
           //Erase the remaining element
           #INO_tMergeBuffer.rgtMessages[#INO_tMergeBuffer.dNumOfMessage - 1].dCodeEvent := 0;
           #INO_tMergeBuffer.rgtMessages[#INO_tMergeBuffer.dNumOfMessage - 1].strIdent := '';
           #INO_tMergeBuffer.rgtMessages[#INO_tMergeBuffer.dNumOfMessage - 1].dEvent1 := 0;
           #INO_tMergeBuffer.rgtMessages[#INO_tMergeBuffer.dNumOfMessage - 1].dEvent2 := 0;
           #INO_tMergeBuffer.rgtMessages[#INO_tMergeBuffer.dNumOfMessage - 1].dEvent3 := 0;
           #INO_tMergeBuffer.rgtMessages[#INO_tMergeBuffer.dNumOfMessage - 1].dEvent4 := 0;
           #INO_tMergeBuffer.rgtMessages[#INO_tMergeBuffer.dNumOfMessage - 1].dEvent5 := 0;
           #INO_tMergeBuffer.rgtMessages[#INO_tMergeBuffer.dNumOfMessage - 1].dEvent6 := 0;
           #INO_tMergeBuffer.rgtMessages[#INO_tMergeBuffer.dNumOfMessage - 1].dEvent7 := 0;
           #INO_tMergeBuffer.rgtMessages[#INO_tMergeBuffer.dNumOfMessage - 1].dEvent8 := 0;
           #INO_tMergeBuffer.rgtMessages[#INO_tMergeBuffer.dNumOfMessage - 1].dEvent9 := 0;
           #INO_tMergeBuffer.rgtMessages[#INO_tMergeBuffer.dNumOfMessage - 1].dEvent10 := 0;

           //Decrement the counter
           //
           #INO_tMergeBuffer.dNumOfMessage := #INO_tMergeBuffer.dNumOfMessage - 1;

       END_IF;


       #OUT_xDataAvailable := true;


   END_IF;
END_FUNCTION

// folder: 06_Output

FUNCTION "OutputTaskSlow" : Void   // FC11, LAD
{ S7_Optimized_Access := 'TRUE' }
VERSION : 0.1
   VAR_TEMP
      TMP_xSpareOFF : Bool;
   END_VAR
BEGIN

REGION Network 1 (SCL)
   #TMP_xSpareOFF := FALSE;


   "o.R195AP1.R251KA1.EncoderCommutation" :="FB_DigitizerManager_V1_00_IDB".OUTPUTS.xSelectEncoder1;
   "o.R195AP1.R251KA2.Jog" := "FB_DigitizerManager_V1_00_IDB".OUTPUTS.xEnableJog;
   "o.R195AP1.R252HL1.SafetiesON" :="Z200".tOutputs.xSafetiesON;

   "o.R195AP1.R251KA3.CpuASerSel":="Z200".tOutputs.xPLC1On;
   "o.R195AP1.R251KA4.CpuBSerSel" := "Z200".tOutputs.xPLC2On;

   "o.R195AP1.R252HL2.EnableCPUA" :="Z200".tOutputs.xPLC1On;
   "o.R195AP1.R252HL2.EnableCPUB" :="Z200".tOutputs.xPLC2On;


   "o.MCC1256B1_IDevice" := "FB_YCuts1_V1_00_IDB".OUT_tIDeviceData;
   "o.MCC1256B2_IDevice" := "FB_YCuts2_V1_00_IDB".OUT_tIDeviceData;


   "o.MCC1204_IDeviceToMarkers" := "FB_Markers_V1.00_IDB".OUT_tIDeviceData;

   "o.R195AP1.M216YV1.DigitizerRise/descentEncoder1" := "FB_Digitizer_1_V1_00_IDB".OUTPUTS.xDescentEncoder;
   "o.R195AP1.M216YV2.DigitizeRise/descentEncoder2" := "FB_Digitizer_2_V1_00_IDB".OUTPUTS.xDescentEncoder;
   "o.R195AP1.R429YV1.StartFillingPumpCuttingTank" := "FB_Oil_V1_00_IDB".OUTPUT.xTankFillCut;
   "o.R195AP1.M221YV2.UpperHolderControl" := "FB_Snaproll_V1_00_IDB".tOutputs.xContrastActivation;
   "o.R195AP1.M221YV1.BreakoutBarControl" := "FB_Snaproll_V1_00_IDB".tOutputs.xRiseSnap;

   "o.R195AP1.M221HL1.CutTrasversalBridge1" := "FB_Snaproll_V1_00_IDB".tOutputs.rgxHLCutDoneXC[0];
   "o.R195AP1.M221HL2.CutTrasversalBridge2" := "FB_Snaproll_V1_00_IDB".tOutputs.rgxHLCutDoneXC[1];
   "o.R195AP1.M221HL3.CutTrasversalBridge3" := "FB_Snaproll_V1_00_IDB".tOutputs.rgxHLCutDoneXC[2];


   "o.R195AP1.M212SB3.M212SB6.GlassRequestQlt" := "FB_ManInsp_V1_00_IDB".OUTPUT.rgxQualityButtonsLamp[0];






   "o_HSCOutput_Count2".swGate := "FB_Digitizer_1_V1_00_IDB".OUTPUTS.xCounterSWGate;
   "o_HSCOutput_Count3".swGate := "FB_Digitizer_2_V1_00_IDB".OUTPUTS.xCounterSWGate;
END_REGION
END_FUNCTION

FUNCTION "OutputTaskFast" : Void   // FC12, LAD
{ S7_Optimized_Access := 'TRUE' }
VERSION : 0.1
BEGIN

REGION Network 1 (SCL)
   "o.R195AP1.R252KA1.SCANNER.RiseBreakingBar" := "FB_ISRASNAP_V1_00_IDB".tOutputs.xSnap;
   "o.R195AP1.R252KA2.SCANNER.GlassToSQC" := "FB_ISRASNAP_V1_00_IDB".tOutputs.xSnapQlt;
   "o.R195AP1.A252KA3.SCANNER.NoGlassBreak" := "FB_ISRA5D_IDB".OUT_xGlassBreak;

   "o_HSCOutput_Count1" := "FB_TrackEncoder_V1_00_IDB".OUT_tHSCCount;
END_REGION
END_FUNCTION

FUNCTION "OutputTaskMedium" : Void   // FC13, LAD
{ S7_Optimized_Access := 'TRUE' }
VERSION : 0.1
BEGIN
END_FUNCTION

FUNCTION "Output_Z201_Idevice" : Void   // FC31, LAD
{ S7_Optimized_Access := 'TRUE' }
VERSION : 0.1
   VAR_TEMP
      TMP_xSpareOFF : Bool;
   END_VAR
BEGIN

REGION Network 1 (SCL)
   #TMP_xSpareOFF := FALSE;



   "FB_CommunicationZ300_V1.00_DB".OUT.Z200.tOUT_Mcc1201."xA47.7" := "Z201".tOutputs.xSafetiesON;

   "FB_CommunicationZ300_V1.00_DB".OUT.Z200.tOUT_Mcc1301."xE.A126.0" := "Z201".tOutputs.xHLResetAnomaly;

   //"o.CS4202.E406AP1.E547SB3.StartCleaningZ301" := "Check";
   //"o.CS4202.E406AP1.E547SB2.ResetAnomalyZ301" := "Check";
   //"o.CS4202.E406AP1.E547SB2.ResetAnomalyZ302" := "Check";
   //"o.CS4202.E406AP1.E547SB4.StopCleaningZ301" := "Check";

   "FB_CommunicationZ300_V1.00_DB".OUT.Z200.tOUT_Mcc1301."xE.A126.6" := "FB_BD_BreakPH_V1_00_IDB".OUTPUT.xSirenBreakAlarm OR"FB_BD_DigitizerPH_V1_00_IDB".OUTPUT.xSirenBreakAlarm ;
   "FB_CommunicationZ300_V1.00_DB".OUT.Z200.tOUT_Mcc1201."xA46.0" :=  "FB_BD_BreakPH_V1_00_IDB".OUTPUT.xLampBreakAlarm OR  "FB_BD_DigitizerPH_V1_00_IDB".OUTPUT.xLampBreakAlarm;


   "FB_CommunicationZ300_V1.00_DB".OUT.Z200.tOUT_Mcc1201."xA87.2" := "FB_DropConveyor_IDB".OUTPUT.xDescentDrop;
   "FB_CommunicationZ300_V1.00_DB".OUT.Z200.tOUT_Mcc1201."xA87.1" := "FB_DropConveyor_IDB".OUTPUT.xRiseDrop;
   "FB_CommunicationZ300_V1.00_DB".OUT.Z200.tOUT_Mcc1201."xA44.4" := true;
   "FB_CommunicationZ300_V1.00_DB".OUT.Z200.tOUT_Mcc1201."xA46.3" := "FB_DropConveyor_IDB".OUTPUT.xHLDoorOpen;
   "FB_CommunicationZ300_V1.00_DB".OUT.Z200.tOUT_Mcc1201."xA46.2" := "FB_DropConveyor_IDB".OUTPUT.xHLUpDownPushbutton;
   "FB_CommunicationZ300_V1.00_DB".OUT.Z200.tOUT_Mcc1201."xA46.5":= "FB_DropConveyor_IDB".OUTPUT.xHLDoorOpen;
   "FB_CommunicationZ300_V1.00_DB".OUT.Z200.tOUT_Mcc1201."xA46.6" := "FB_DropConveyor_IDB".OUTPUT.xHLUpDownPushbutton;

   "FB_CommunicationZ300_V1.00_DB".OUT.Z200.tOUT_Mcc1201."xA87.4" := "FB_BreakerM206_V1_00_IDB".OUTPUT.xBreakerRun;
   "FB_CommunicationZ300_V1.00_DB".OUT.Z200.tOUT_Mcc1201."xA44.0" := "FB_BreakerM206_V1_00_IDB".OUTPUT.xToScrapingUnderZ200;

   "FB_CommunicationZ300_V1.00_DB".OUT.Z200.tOUT_Mcc1201."xA86.0":="Z201".tOutputs.xRunFanM216;
   "FB_CommunicationZ300_V1.00_DB".OUT.Z200.tOUT_Mcc1201."xA87.6" := "Z201".tOutputs.xRunFanM209;
   "FB_CommunicationZ300_V1.00_DB".OUT.Z200.tOUT_Mcc1201."xA47.0" := "Z201".tOutputs.xHLchipBlowerM209On;

   "FB_CommunicationZ300_V1.00_DB".OUT.Z200.tOUT_Mcc1201."xA47.2" := "FB_BreakerM206_V1_00_IDB".OUTPUT.xHlScrapinglineReady;
   "FB_CommunicationZ300_V1.00_DB".OUT.Z200.tOUT_Mcc1201."xA47.3" := "FB_BreakerM206_V1_00_IDB".OUTPUT.xHlScrapinglineNotReady;
   "FB_CommunicationZ300_V1.00_DB".OUT.Z200.tOUT_Mcc1201."xA44.3" := "Z201".tOutputs.xHAAlarm;

   "FB_CommunicationZ300_V1.00_DB".OUT.Z200.tOUT_Mcc1201."xA45.0" := "FB_IO_EmergencyCuttingBridge_DB".OUT_xSnap;
   "FB_CommunicationZ300_V1.00_DB".OUT.Z200.tOUT_Mcc1201."xA45.3" := "FB_IO_EmergencyCuttingBridge_DB".OUT_xStartCutCycle;
END_REGION
END_FUNCTION

// folder: 07_ArrayScada

FUNCTION "SCADA_Mapping" : Void   // FC26, SCL
{ S7_Optimized_Access := 'TRUE' }
VERSION : 0.1
   VAR_TEMP
      TMP_dIndex : DInt;
   END_VAR
BEGIN


       //Move M201 HMR
       "DB_Conveyor_M201_HMI".tHMR.xManualCommandEnabled := "FB_Z200Conveyor_M201_IDB".tHMR.xManualCommandEnabled;
       "DB_Conveyor_M201_HMI".tHMR.dState := "FB_Z200Conveyor_M201_IDB".tHMR.dState;
       "DB_Conveyor_M201_HMI".tHMR.dSpeedFeedback := "FB_Z200Conveyor_M201_IDB".tHMR.dSpeedFeedback;
       "DB_Conveyor_M201_HMI".tHMR.tManCmd.xFdbkRunFw := "FB_Z200Conveyor_M201_IDB".tHMR.tManCmd.xFdbkRunFw;

       //Move M201 HMW
       "FB_Z200Conveyor_M201_IDB".tHMW.xEnableManualCommand := "DB_Conveyor_M201_HMI".tHMW.xEnableManualCommand;
       "FB_Z200Conveyor_M201_IDB".tHMW.tManCmd.xRunFw := "DB_Conveyor_M201_HMI".tHMW.tManCmd.xRunFw;
       "FB_Z200Conveyor_M201_IDB".tHMW.dCurrentLimit := "DB_Conveyor_M201_HMI".tHMW.dCurrentLimit;
       "FB_Z200Conveyor_M201_IDB".tHMW.dSpeedCorrection := "DB_Conveyor_M201_HMI".tHMW.dSpeedCorrection;

       //Move M201 ALM
       "DB_Conveyor_M201_HMI".tALM.tF :="FB_Z200Conveyor_M201_IDB".tALM.tF;
       "DB_Conveyor_M201_HMI".tALM.tS := "FB_Z200Conveyor_M201_IDB".tALM.tS;
       "DB_Conveyor_M201_HMI".tALM.tW := "FB_Z200Conveyor_M201_IDB".tALM.tW;

       //Move M204 HMR
       "DB_Conveyor_M204_HMI".tHMR.xManualCommandEnabled := "FB_Z200Conveyor_M204_IDB".tHMR.xManualCommandEnabled;
       "DB_Conveyor_M204_HMI".tHMR.dState := "FB_Z200Conveyor_M204_IDB".tHMR.dState;
       "DB_Conveyor_M204_HMI".tHMR.dSpeedFeedback := "FB_Z200Conveyor_M204_IDB".tHMR.dSpeedFeedback;
       "DB_Conveyor_M204_HMI".tHMR.tManCmd.xFdbkRunFw := "FB_Z200Conveyor_M204_IDB".tHMR.tManCmd.xFdbkRunFw;

       //Move M204 HMW
       "FB_Z200Conveyor_M204_IDB".tHMW.xEnableManualCommand := "DB_Conveyor_M204_HMI".tHMW.xEnableManualCommand;
       "FB_Z200Conveyor_M204_IDB".tHMW.tManCmd.xRunFw := "DB_Conveyor_M204_HMI".tHMW.tManCmd.xRunFw;
       "FB_Z200Conveyor_M204_IDB".tHMW.dCurrentLimit := "DB_Conveyor_M204_HMI".tHMW.dCurrentLimit;
       "FB_Z200Conveyor_M204_IDB".tHMW.dSpeedCorrection := "DB_Conveyor_M204_HMI".tHMW.dSpeedCorrection;

       //Move M204 ALM
       "DB_Conveyor_M204_HMI".tALM.tF := "FB_Z200Conveyor_M204_IDB".tALM.tF;
       "DB_Conveyor_M204_HMI".tALM.tS := "FB_Z200Conveyor_M204_IDB".tALM.tS;
       "DB_Conveyor_M204_HMI".tALM.tW := "FB_Z200Conveyor_M204_IDB".tALM.tW;

       //Move M205 HMR
       "DB_Conveyor_M205_HMI".tHMR.xManualCommandEnabled := "FB_Z200Conveyor_M205_IDB".tHMR.xManualCommandEnabled;
       "DB_Conveyor_M205_HMI".tHMR.dState := "FB_Z200Conveyor_M205_IDB".tHMR.dState;
       "DB_Conveyor_M205_HMI".tHMR.dSpeedFeedback := "FB_Z200Conveyor_M205_IDB".tHMR.dSpeedFeedback;
       "DB_Conveyor_M205_HMI".tHMR.tManCmd.xFdbkRunFw := "FB_Z200Conveyor_M205_IDB".tHMR.tManCmd.xFdbkRunFw;

       //Move M205 HMW
       "FB_Z200Conveyor_M205_IDB".tHMW.xEnableManualCommand := "DB_Conveyor_M205_HMI".tHMW.xEnableManualCommand;
       "FB_Z200Conveyor_M205_IDB".tHMW.tManCmd.xRunFw := "DB_Conveyor_M205_HMI".tHMW.tManCmd.xRunFw;
       "FB_Z200Conveyor_M205_IDB".tHMW.dCurrentLimit := "DB_Conveyor_M205_HMI".tHMW.dCurrentLimit;
       "FB_Z200Conveyor_M205_IDB".tHMW.dSpeedCorrection := "DB_Conveyor_M205_HMI".tHMW.dSpeedCorrection;

       //Move M205 ALM
       "DB_Conveyor_M205_HMI".tALM.tF := "FB_Z200Conveyor_M205_IDB".tALM.tF;


       //Move M208 HMR
       "DB_Conveyor_M208_HMI".tHMR.xManualCommandEnabled := "FB_Z200Conveyor_M208_IDB".tHMR.xManualCommandEnabled;
       "DB_Conveyor_M208_HMI".tHMR.dState := "FB_Z200Conveyor_M208_IDB".tHMR.dState;
       "DB_Conveyor_M208_HMI".tHMR.dSpeedFeedback := "FB_Z200Conveyor_M208_IDB".tHMR.dSpeedFeedback;
       "DB_Conveyor_M208_HMI".tHMR.tManCmd.xFdbkRunFw := "FB_Z200Conveyor_M208_IDB".tHMR.tManCmd.xFdbkRunFw;

       //Move M208 HMW
       "FB_Z200Conveyor_M208_IDB".tHMW.xEnableManualCommand := "DB_Conveyor_M208_HMI".tHMW.xEnableManualCommand;
       "FB_Z200Conveyor_M208_IDB".tHMW.tManCmd.xRunFw := "DB_Conveyor_M208_HMI".tHMW.tManCmd.xRunFw;
       "FB_Z200Conveyor_M208_IDB".tHMW.dCurrentLimit := "DB_Conveyor_M208_HMI".tHMW.dCurrentLimit;
       "FB_Z200Conveyor_M208_IDB".tHMW.dSpeedCorrection := "DB_Conveyor_M208_HMI".tHMW.dSpeedCorrection;

       //Move M208 ALM
       "DB_Conveyor_M208_HMI".tALM.tF := "FB_Z200Conveyor_M208_IDB".tALM.tF;
       "DB_Conveyor_M208_HMI".tALM.tS:= "FB_Z200Conveyor_M208_IDB".tALM.tS;
       "DB_Conveyor_M208_HMI".tALM.tW := "FB_Z200Conveyor_M208_IDB".tALM.tW;

        //Move M211 HMR
       "DB_Conveyor_M211_HMI".tHMR.xManualCommandEnabled := "FB_Z200Conveyor_M211_iDB".tHMR.xManualCommandEnabled;
       "DB_Conveyor_M211_HMI".tHMR.dState := "FB_Z200Conveyor_M211_iDB".tHMR.dState;
       "DB_Conveyor_M211_HMI".tHMR.dSpeedFeedback := "FB_Z200Conveyor_M211_iDB".tHMR.dSpeedFeedback;
       "DB_Conveyor_M211_HMI".tHMR.tManCmd.xFdbkRunFw := "FB_Z200Conveyor_M211_iDB".tHMR.tManCmd.xFdbkRunFw;

       //Move M211 HMW
       "FB_Z200Conveyor_M211_iDB".tHMW.xEnableManualCommand := "DB_Conveyor_M211_HMI".tHMW.xEnableManualCommand;
       "FB_Z200Conveyor_M211_iDB".tHMW.tManCmd.xRunFw := "DB_Conveyor_M211_HMI".tHMW.tManCmd.xRunFw;
       "FB_Z200Conveyor_M211_iDB".tHMW.dCurrentLimit := "DB_Conveyor_M211_HMI".tHMW.dCurrentLimit;
       "FB_Z200Conveyor_M211_iDB".tHMW.dSpeedCorrection := "DB_Conveyor_M211_HMI".tHMW.dSpeedCorrection;

       //Move M211 ALM
       "DB_Conveyor_M211_HMI".tALM.tF := "FB_Z200Conveyor_M211_iDB".tALM.tF;
       "DB_Conveyor_M211_HMI".tALM.tS := "FB_Z200Conveyor_M211_iDB".tALM.tS;
       "DB_Conveyor_M211_HMI".tALM.tW := "FB_Z200Conveyor_M211_iDB".tALM.tW;



       //Move M214 HMR
       "DB_Conveyor_M214_HMI".tHMR.xManualCommandEnabled := "FB_Z200Conveyor_M214_iDB".tHMR.xManualCommandEnabled;
       "DB_Conveyor_M214_HMI".tHMR.dState := "FB_Z200Conveyor_M214_iDB".tHMR.dState;
       "DB_Conveyor_M214_HMI".tHMR.dSpeedFeedback := "FB_Z200Conveyor_M214_iDB".tHMR.dSpeedFeedback;
       "DB_Conveyor_M214_HMI".tHMR.tManCmd.xFdbkRunFw := "FB_Z200Conveyor_M214_iDB".tHMR.tManCmd.xFdbkRunFw;

       //Move M214 HMW
       "FB_Z200Conveyor_M214_iDB".tHMW.xEnableManualCommand := "DB_Conveyor_M214_HMI".tHMW.xEnableManualCommand;
       "FB_Z200Conveyor_M214_iDB".tHMW.tManCmd.xRunFw := "DB_Conveyor_M214_HMI".tHMW.tManCmd.xRunFw;
       "FB_Z200Conveyor_M214_iDB".tHMW.dCurrentLimit := "DB_Conveyor_M214_HMI".tHMW.dCurrentLimit;
       "FB_Z200Conveyor_M214_iDB".tHMW.dSpeedCorrection := "DB_Conveyor_M214_HMI".tHMW.dSpeedCorrection;

       //Move M214 ALM
       "DB_Conveyor_M214_HMI".tALM.tF := "FB_Z200Conveyor_M214_iDB".tALM.tF;
       "DB_Conveyor_M214_HMI".tALM.tS := "FB_Z200Conveyor_M214_iDB".tALM.tS;
       "DB_Conveyor_M214_HMI".tALM.tW := "FB_Z200Conveyor_M214_iDB".tALM.tW;

       //Move M218 HMR
       "DB_Conveyor_M218_HMI".tHMR.xManualCommandEnabled := "FB_Z200Conveyor_M218_IDB".tHMR.xManualCommandEnabled;
       "DB_Conveyor_M218_HMI".tHMR.dState := "FB_Z200Conveyor_M218_IDB".tHMR.dState;
       "DB_Conveyor_M218_HMI".tHMR.dSpeedFeedback := "FB_Z200Conveyor_M218_IDB".tHMR.dSpeedFeedback;
       "DB_Conveyor_M218_HMI".tHMR.tManCmd.xFdbkRunFw := "FB_Z200Conveyor_M218_IDB".tHMR.tManCmd.xFdbkRunFw;

       //Move M218 HMW
       "FB_Z200Conveyor_M218_IDB".tHMW.xEnableManualCommand := "DB_Conveyor_M218_HMI".tHMW.xEnableManualCommand;
       "FB_Z200Conveyor_M218_IDB".tHMW.tManCmd.xRunFw := "DB_Conveyor_M218_HMI".tHMW.tManCmd.xRunFw;
       "FB_Z200Conveyor_M218_IDB".tHMW.dCurrentLimit := "DB_Conveyor_M218_HMI".tHMW.dCurrentLimit;
       "FB_Z200Conveyor_M218_IDB".tHMW.dSpeedCorrection := "DB_Conveyor_M218_HMI".tHMW.dSpeedCorrection;

       //Move M218 ALM
       "DB_Conveyor_M218_HMI".tALM.tF := "FB_Z200Conveyor_M218_IDB".tALM.tF;
       "DB_Conveyor_M218_HMI".tALM.tS := "FB_Z200Conveyor_M218_IDB".tALM.tS;
       "DB_Conveyor_M218_HMI".tALM.tW := "FB_Z200Conveyor_M218_IDB".tALM.tW;

       //Move M206 HMR
       "DB_Breaker_M206_HMI".tHMR.xSpare1 :="FB_BreakerM206_V1_00_IDB".tHMR.xEnabledRunAlwaysModeBreaker;
       "DB_Breaker_M206_HMI".tHMR.xManualCommandEnabled := "FB_BreakerM206_V1_00_IDB".tHMR.xManualCommandEnabled;
       "DB_Breaker_M206_HMI".tHMR.tManCmd.xRunFdbk := "FB_BreakerM206_V1_00_IDB".tHMR.tManCmd.xRunFdbk;

       //Move M206 HMW
       "FB_BreakerM206_V1_00_IDB".tHMW.dBreakerRetainTime_s := "DB_Breaker_M206_HMI".tHMW.dBreakerRetainTime_s;
       "FB_BreakerM206_V1_00_IDB".tHMW.xEnableManualCommand := "DB_Breaker_M206_HMI".tHMW.xEnableManualCommand;
       "FB_BreakerM206_V1_00_IDB".tHMW.xEnableRunAlwaysModeBreaker := "DB_Breaker_M206_HMI".tHMW.xEnableRunAlwaysModeBreaker;
       "FB_BreakerM206_V1_00_IDB".tHMW.tManCmd.xRun := "DB_Breaker_M206_HMI".tHMW.tManCmd.xRun;

       //Move M206 ALM 
       "DB_Breaker_M206_HMI".tALM.tF :="FB_BreakerM206_V1_00_IDB".tALM.tF;
       "DB_Breaker_M206_HMI".tALM.tS :="FB_BreakerM206_V1_00_IDB".tALM.tS;
       "DB_Breaker_M206_HMI".tALM.tW :="FB_BreakerM206_V1_00_IDB".tALM.tW;

       //Move MAN INSP HMR
       //
       "DB_MAN_INSP_HMI".tHMR.xManualCommandEnabled := "FB_ManInsp_V1_00_IDB".tHMR.xManComEn;
       "DB_MAN_INSP_HMI".tHMR.dDistanceSnaproll_cmm := "FB_ManInsp_V1_00_IDB".tHMR.dDistanceSnaproll_cmm;
       "DB_MAN_INSP_HMI".tHMR.tManCmd.xSpare1 := "FB_ManInsp_V1_00_IDB".tHMR.tManFdbk.xFanCommand; 

       //Move MAN INSP   HMW
       "FB_ManInsp_V1_00_IDB".tHMW.xUpdateDistanceSnaproll := "DB_MAN_INSP_HMI".tHMW.xUpdateDistanceSnaproll;
       "FB_ManInsp_V1_00_IDB".tHMW.xEnDisManCom := "DB_MAN_INSP_HMI".tHMW.xEnableManualCommand;
       "FB_ManInsp_V1_00_IDB".tHMW.rgxEnabledContinuosDef[0] := "DB_MAN_INSP_HMI".tHMW."xEnabledContinuosDef[0]";
       "FB_ManInsp_V1_00_IDB".tHMW.rgxEnabledContinuosDef[1] := "DB_MAN_INSP_HMI".tHMW."xEnabledContinuosDef[1]";
       "FB_ManInsp_V1_00_IDB".tHMW.rgxEnabledContinuosDef[2] := "DB_MAN_INSP_HMI".tHMW."xEnabledContinuosDef[2]";
       "FB_ManInsp_V1_00_IDB".tHMW.rgxEnabledContinuosDef[3] := "DB_MAN_INSP_HMI".tHMW."xEnabledContinuosDef[3]";
       "FB_ManInsp_V1_00_IDB".tHMW.tMan.xFanCommand := "DB_MAN_INSP_HMI".tHMW.tManCmd.xSpare0;


       //Move MAN INSP  ALM  
       "DB_MAN_INSP_HMI".tALM.tF := "FB_ManInsp_V1_00_IDB".tALM.tF;
       "DB_MAN_INSP_HMI".tALM.tS := "FB_ManInsp_V1_00_IDB".tALM.tS;
       "DB_MAN_INSP_HMI".tALM.tW := "FB_ManInsp_V1_00_IDB".tALM.tW;

       //Move BREAK DETECTOR HMR

       "DB_Break_detector_M202_HMI".tHMR."xPhotoStatus[0]" := "FB_BD_BreakPH_V1_00_IDB".tHMR.rgxPhotoStatus[0];
       "DB_Break_detector_M202_HMI".tHMR."xPhotoStatus[1]" := "FB_BD_BreakPH_V1_00_IDB".tHMR.rgxPhotoStatus[1];
       "DB_Break_detector_M202_HMI".tHMR."xPhotoStatus[2]" := "FB_BD_BreakPH_V1_00_IDB".tHMR.rgxPhotoStatus[2];
       "DB_Break_detector_M202_HMI".tHMR."xPhotoStatus[3]" := "FB_BD_BreakPH_V1_00_IDB".tHMR.rgxPhotoStatus[3];
       "DB_Break_detector_M202_HMI".tHMR."xPhotoStatus[4]" := "FB_BD_BreakPH_V1_00_IDB".tHMR.rgxPhotoStatus[4];
       "DB_Break_detector_M202_HMI".tHMR."xPhotoStatus[5]" := "FB_BD_BreakPH_V1_00_IDB".tHMR.rgxPhotoStatus[5];
       "DB_Break_detector_M202_HMI".tHMR."xPhotoStatus[6]" := "FB_BD_BreakPH_V1_00_IDB".tHMR.rgxPhotoStatus[6];
       "DB_Break_detector_M202_HMI".tHMR."xPhotoStatus[7]" := "FB_BD_BreakPH_V1_00_IDB".tHMR.rgxPhotoStatus[7];
       "DB_Break_detector_M202_HMI".tHMR."xPhotoStatus[8]" := "FB_BD_BreakPH_V1_00_IDB".tHMR.rgxPhotoStatus[8];
       "DB_Break_detector_M202_HMI".tHMR."xPhotoStatus[9]" := "FB_BD_BreakPH_V1_00_IDB".tHMR.rgxPhotoStatus[9];

       "DB_Break_detector_M202_HMI".tHMR.dDistanceSnaproll_cmm := "FB_BD_BreakPH_V1_00_IDB".tHMR.dDistanceSnaproll_cmm;
       "DB_Break_detector_M202_HMI".tHMR.dStatus := "FB_BD_BreakPH_V1_00_IDB".tHMR.dStatus;
       "DB_Break_detector_M202_HMI".tHMR."dPhotoAbilitation[0]" := "FB_BD_BreakPH_V1_00_IDB".tHMR.rgdPhotoAbilitation[0];
       "DB_Break_detector_M202_HMI".tHMR."dPhotoAbilitation[1]" := "FB_BD_BreakPH_V1_00_IDB".tHMR.rgdPhotoAbilitation[1];
       "DB_Break_detector_M202_HMI".tHMR."dPhotoAbilitation[2]" := "FB_BD_BreakPH_V1_00_IDB".tHMR.rgdPhotoAbilitation[2];
       "DB_Break_detector_M202_HMI".tHMR."dPhotoAbilitation[3]" := "FB_BD_BreakPH_V1_00_IDB".tHMR.rgdPhotoAbilitation[3];
       "DB_Break_detector_M202_HMI".tHMR."dPhotoAbilitation[4]" := "FB_BD_BreakPH_V1_00_IDB".tHMR.rgdPhotoAbilitation[4];
       "DB_Break_detector_M202_HMI".tHMR."dPhotoAbilitation[5]" := "FB_BD_BreakPH_V1_00_IDB".tHMR.rgdPhotoAbilitation[5];
       "DB_Break_detector_M202_HMI".tHMR."dPhotoAbilitation[6]" := "FB_BD_BreakPH_V1_00_IDB".tHMR.rgdPhotoAbilitation[6];
       "DB_Break_detector_M202_HMI".tHMR."dPhotoAbilitation[7]" := "FB_BD_BreakPH_V1_00_IDB".tHMR.rgdPhotoAbilitation[7];
       "DB_Break_detector_M202_HMI".tHMR."dPhotoAbilitation[8]" := "FB_BD_BreakPH_V1_00_IDB".tHMR.rgdPhotoAbilitation[8];
       "DB_Break_detector_M202_HMI".tHMR."dPhotoAbilitation[9]" := "FB_BD_BreakPH_V1_00_IDB".tHMR.rgdPhotoAbilitation[9];

       //Move BREAK DETECTOR HMW
       "FB_BD_BreakPH_V1_00_IDB".tHMW.xUpdateDistanceSnap := "DB_Break_detector_M202_HMI".tHMW.xUpdateDistanceSnaproll;

       "FB_BD_BreakPH_V1_00_IDB".tHMW.rgxEnabledPhotocell[0] := "DB_Break_detector_M202_HMI".tHMW."xPhotoEnabled[0]";
       "FB_BD_BreakPH_V1_00_IDB".tHMW.rgxEnabledPhotocell[1] := "DB_Break_detector_M202_HMI".tHMW."xPhotoEnabled[1]";
       "FB_BD_BreakPH_V1_00_IDB".tHMW.rgxEnabledPhotocell[2] := "DB_Break_detector_M202_HMI".tHMW."xPhotoEnabled[2]";
       "FB_BD_BreakPH_V1_00_IDB".tHMW.rgxEnabledPhotocell[3] := "DB_Break_detector_M202_HMI".tHMW."xPhotoEnabled[3]";
       "FB_BD_BreakPH_V1_00_IDB".tHMW.rgxEnabledPhotocell[4] := "DB_Break_detector_M202_HMI".tHMW."xPhotoEnabled[4]";
       "FB_BD_BreakPH_V1_00_IDB".tHMW.rgxEnabledPhotocell[5] := "DB_Break_detector_M202_HMI".tHMW."xPhotoEnabled[5]";
       "FB_BD_BreakPH_V1_00_IDB".tHMW.rgxEnabledPhotocell[6] := "DB_Break_detector_M202_HMI".tHMW."xPhotoEnabled[6]";
       "FB_BD_BreakPH_V1_00_IDB".tHMW.rgxEnabledPhotocell[7] := "DB_Break_detector_M202_HMI".tHMW."xPhotoEnabled[7]";
       "FB_BD_BreakPH_V1_00_IDB".tHMW.rgxEnabledPhotocell[8] := "DB_Break_detector_M202_HMI".tHMW."xPhotoEnabled[8]";
       "FB_BD_BreakPH_V1_00_IDB".tHMW.rgxEnabledPhotocell[9] := "DB_Break_detector_M202_HMI".tHMW."xPhotoEnabled[9]";

       "FB_BD_BreakPH_V1_00_IDB".tHMW.dDistanceSnaproll_cmm := "DB_Break_detector_M202_HMI".tHMW.dDistanceSnaproll_cmm;
       "FB_BD_BreakPH_V1_00_IDB".tHMW.dMinBreakSize_cmm :="DB_Break_detector_M202_HMI".tHMW.dMinBreakSize_cmm;

       //Move BREAK DETECTOR ALM
       "DB_Break_detector_M202_HMI".tALM.tF := "FB_BD_BreakPH_V1_00_IDB".tALM.tF;
       "DB_Break_detector_M202_HMI".tALM.tS := "FB_BD_BreakPH_V1_00_IDB".tALM.tS;
       "DB_Break_detector_M202_HMI".tALM.tW := "FB_BD_BreakPH_V1_00_IDB".tALM.tW;

       //Move ISRA HMR
       "DB_ISRA_HMI".tHMR.xScannerON := "FB_ISRA5D_IDB".tHMR.xScannerON;

       "DB_ISRA_HMI".tHMR.dCurrentGrossWander_cmm := "FB_ISRA5D_IDB".tHMR.dCurrentGrossWander_cmm;
       "DB_ISRA_HMI".tHMR.dCurrentGrossWidth_cmm := "FB_ISRA5D_IDB".tHMR.dCurrentGrossWidth_cmm;
       "DB_ISRA_HMI".tHMR.dCurrentNetWander_cmm := "FB_ISRA5D_IDB".tHMR.dCurrentNetWander_cmm;
       "DB_ISRA_HMI".tHMR.dCurrentNetWidth_cmm := "FB_ISRA5D_IDB".tHMR.dCurrentNetWidth_cmm;
       "DB_ISRA_HMI".tHMR.dDistanceSnaproll_cmm := "FB_ISRA5D_IDB".tHMR.dDistSnapRoll_cmm;
       "DB_ISRA_HMI".tHMR.dDistCenterLine_cmm := "FB_ISRA5D_IDB".tHMR.dDistCenterLine_cmm;
       "DB_ISRA_HMI".tHMR.dInspectionStatus := "FB_ISRA5D_IDB".tHMR.dInspectionStatus;

       //Move ISRA  HMW
       "FB_ISRA5D_IDB".tHMW.xAutoInspEnabled := "DB_ISRA_HMI".tHMW.xAutoInspEnabled;
       "FB_ISRA5D_IDB".tHMW.xUpdDistSnaproll := "DB_ISRA_HMI".tHMW.xUpdateDistanceSnaproll;
       "FB_ISRA5D_IDB".tHMW .xUpdDistCenterLine :="DB_ISRA_HMI".tHMW.xUpdDistCenterLine;
       "FB_ISRA5D_IDB".tHMW .xCalibPosition:= "DB_ISRA_HMI".tHMW.xDefectPositionCalibration;

       "FB_ISRA5D_IDB".tHMW.dDistSnapRoll_cmm := "DB_ISRA_HMI".tHMW.dDistanceSnaproll_cmm;
       "FB_ISRA5D_IDB".tHMW.dDistCenterLine_cmm := "DB_ISRA_HMI".tHMW.dDistCenterLine_cmm;
       "FB_ISRA5D_IDB".tHMW.dCalibDefRealXPos_cmm := "DB_ISRA_HMI".tHMW.dCalibDefectRealPosX_cmm;
       "FB_ISRA5D_IDB".tHMW.dCalibDefRealYPos_cmm := "DB_ISRA_HMI".tHMW.dCalibDefRealYPos_cmm;
       "FB_ISRA5D_IDB".tHMW.dCalibDefTeoXPos_cmm := "DB_ISRA_HMI".tHMW.dCalibDefectTheoPosX_cmm;
       "FB_ISRA5D_IDB".tHMW.dCalibDefTeoYPos_cmm := "DB_ISRA_HMI".tHMW.dCalibDefTeoYPos_cmm;

       //Move ISRA ALM  
       "DB_ISRA_HMI".tALM.tF := "FB_ISRA5D_IDB".tALM.tF;
       "DB_ISRA_HMI".tALM.tS := "FB_ISRA5D_IDB".tALM.tS;
       "DB_ISRA_HMI".tALM.tW := "FB_ISRA5D_IDB".tALM.tW;

       //Move WANDER CAMERA HMR
       "DB_WANDER_HMI".tHMR.dCameraStatus := "FB_WanderCamera_V1_00_IDB".tHMR.dCameraStatus;
       "DB_WANDER_HMI".tHMR.dCurrentGrossWander_cmm := "FB_WanderCamera_V1_00_IDB".tHMR.dCurrentGrossWander_cmm;
       "DB_WANDER_HMI".tHMR.dCurrentGrossWidth_cmm := "FB_WanderCamera_V1_00_IDB".tHMR.dCurrentGrossWidth_cmm;
       "DB_WANDER_HMI".tHMR.dCurrentNetWander_cmm := "FB_WanderCamera_V1_00_IDB".tHMR.dCurrentNetWander_cmm;
       "DB_WANDER_HMI".tHMR.dCurrentNetWidth_cmm := "FB_WanderCamera_V1_00_IDB".tHMR.dCurrentNetWidth_cmm;
       "DB_WANDER_HMI".tHMR.dDistanceSnaproll_cmm := "FB_WanderCamera_V1_00_IDB".tHMR.dDistanceFromSnaproll_cmm;

       //Move WANDER CAMERA HMW
       "FB_WanderCamera_V1_00_IDB".tHMW.xUpdateDistanceFromSnaproll := "DB_WANDER_HMI".tHMW.xUpdateDistanceSnaproll;
       "FB_WanderCamera_V1_00_IDB".tHMW.dDistanceFromSnaproll_cmm := "DB_WANDER_HMI".tHMW.dDistanceSnaproll_cmm;

       //Move WANDER CAMERA ALM  
       "DB_WANDER_HMI".tALM.tF := "FB_WanderCamera_V1_00_IDB".tALM.tF;
       "DB_WANDER_HMI".tALM.tS := "FB_WanderCamera_V1_00_IDB".tALM.tS;
       "DB_WANDER_HMI".tALM.tW := "FB_WanderCamera_V1_00_IDB".tALM.tW;

       //Move M204 HMR
       "DB_Dropconveyor_M204_HMI".tHMR.xUpPosition := "FB_DropConveyor_IDB".tHMR.xUpPosition;
       "DB_Dropconveyor_M204_HMI".tHMR.xDownPosition := "FB_DropConveyor_IDB".tHMR.xDownPosition;

       "DB_Dropconveyor_M204_HMI".tHMR.dDistanceSnaproll_cmm := "FB_DropConveyor_IDB".tHMR.dDistanceFromSnaproll_cmm;
       "DB_Dropconveyor_M204_HMI".tHMR.dMode := "FB_DropConveyor_IDB".tHMR.dMode;
       "DB_Dropconveyor_M204_HMI".tHMR.dStatus := "FB_DropConveyor_IDB".tHMR.dStatus;

       "DB_Dropconveyor_M204_HMI".tHMR.tManCmd.xDescentFdbk := "FB_DropConveyor_IDB".tHMR.tManCmd.xDescentFdbk;
       "DB_Dropconveyor_M204_HMI".tHMR.tManCmd.xRiseFdbk := "FB_DropConveyor_IDB".tHMR.tManCmd.xRiseFdbk;

       //Move M204 HMW
       "FB_DropConveyor_IDB".tHMW.xEnabledBreakingDetection := "DB_Dropconveyor_M204_HMI".tHMW.xEnabledBreakingDetection;
       "FB_DropConveyor_IDB".tHMW.xForceDown := "DB_Dropconveyor_M204_HMI".tHMW.xForceDown;
       "FB_DropConveyor_IDB".tHMW.xForceUp := "DB_Dropconveyor_M204_HMI".tHMW.xForceUp;
       "FB_DropConveyor_IDB".tHMW.xRequestDown := "DB_Dropconveyor_M204_HMI".tHMW.xRequestDown;
       "FB_DropConveyor_IDB".tHMW.xRequestUp := "DB_Dropconveyor_M204_HMI".tHMW.xRequestUp;
       "FB_DropConveyor_IDB".tHMW.xUpdateDistanceFromSnaproll := "DB_Dropconveyor_M204_HMI".tHMW.xUpdateDistanceSnaproll;

       "FB_DropConveyor_IDB".tHMW.tManCmd.xDescent := "DB_Dropconveyor_M204_HMI".tHMW.tManCmd.xDescent;
       "FB_DropConveyor_IDB".tHMW.tManCmd.xRise := "DB_Dropconveyor_M204_HMI".tHMW.tManCmd.xRise;

       "FB_DropConveyor_IDB".tHMW.dDistanceFromSnaproll_cmm := "DB_Dropconveyor_M204_HMI".tHMW.dDistanceSnaproll_cmm;

       //Move M204 ALM 
       "DB_Dropconveyor_M204_HMI".tALM.tF := "FB_DropConveyor_IDB".tALM.tF;
       "DB_Dropconveyor_M204_HMI".tALM.tS := "FB_DropConveyor_IDB".tALM.tS;
       "DB_Dropconveyor_M204_HMI".tALM.tW := "FB_DropConveyor_IDB".tALM.tW;

       //Move BPS_A ALM
       "DB_BPS_A_HMI".tALM.tF := "FB_BPSEthLink_ServerA_V1_00_IDB".tALM.tF;
       "DB_BPS_A_HMI".tALM.tS := "FB_BPSEthLink_ServerA_V1_00_IDB".tALM.tS;
       "DB_BPS_A_HMI".tALM.tW := "FB_BPSEthLink_ServerA_V1_00_IDB".tALM.tW;

       //Move BPS_B ALM
       "DB_BPS_B_HMI".tALM.tF := "FB_BPSEthLink_ServerB_V1_00_IDB".tALM.tF;
       "DB_BPS_B_HMI".tALM.tS := "FB_BPSEthLink_ServerB_V1_00_IDB".tALM.tS;
       "DB_BPS_B_HMI".tALM.tW := "FB_BPSEthLink_ServerB_V1_00_IDB".tALM.tW;

       //Move OIL HMR
       "DB_Oil_Manager_HMI".tHMR.xManualCommandEnabled := "FB_Oil_V1_00_IDB".tHMR.xManComEn;
       "DB_Oil_Manager_HMI".tHMR.xOilAtMax := "FB_Oil_V1_00_IDB".tHMR.xOilAtMax;
       "DB_Oil_Manager_HMI".tHMR.xOilAtMin := "FB_Oil_V1_00_IDB".tHMR.xOilAtMin;

       "DB_Oil_Manager_HMI".tHMR.tManCmd.xFillTank := "FB_Oil_V1_00_IDB".tHMR.tManFdbk.xFillTank;

       "DB_Oil_Manager_HMI".tHMR.dStatus := "FB_Oil_V1_00_IDB".tHMR.dStatus;

       //Move OIL  HMW
       "FB_Oil_V1_00_IDB".tHMW.xEnDisManCom := "DB_Oil_Manager_HMI".tHMW.xEnableManualCommand;

       "FB_Oil_V1_00_IDB".tHMW.tMan.xFillTank := "DB_Oil_Manager_HMI".tHMW.tManCmd.xFillTank;

       //Move OIL ALM  
       "DB_Oil_Manager_HMI".tALM.tF := "FB_Oil_V1_00_IDB".tALM.tF;
       "DB_Oil_Manager_HMI".tALM.tS := "FB_Oil_V1_00_IDB".tALM.tS;
       "DB_Oil_Manager_HMI".tALM.tW := "FB_Oil_V1_00_IDB".tALM.tW;

       //Move LEHR SPEED HMR
       "DB_Lehr_Speed_HMI".tHMR.dActualSpeedSource := "FB_LehrSpeed_IDB".tHMR.dActualSpeedSource;
       "DB_Lehr_Speed_HMI".tHMR.dActualSpeedValue_mm_min := "FB_LehrSpeed_IDB".tHMR.dActualSpeedValue_mm_min;
       "DB_Lehr_Speed_HMI".tHMR.dEncoder1Status := "FB_LehrSpeed_IDB".tHMR.dEncoder1Status;
       "DB_Lehr_Speed_HMI".tHMR.dActualSpeedValueToConveyor_mm_min := "FB_LehrSpeed_IDB".tHMR.dActualSpeedValueToConveyor_mm_min;
       "DB_Lehr_Speed_HMI".tHMR.dEncoder2Status := "FB_LehrSpeed_IDB".tHMR.dEncoder2Status;
       "DB_Lehr_Speed_HMI".tHMR.dEncoder1Value_mm_min := "FB_LehrSpeed_IDB".tHMR.dEncoder1Value_mm_min;
       "DB_Lehr_Speed_HMI".tHMR.dEncoder2Value_mm_min := "FB_LehrSpeed_IDB".tHMR.dEncoder2Value_mm_min;
       "DB_Lehr_Speed_HMI".tHMR.dEthStatus := "FB_LehrSpeed_IDB".tHMR.dEthStatus;
       "DB_Lehr_Speed_HMI".tHMR.dEthValue_mm_min := "FB_LehrSpeed_IDB".tHMR.dEthValue_mm_min;
       "DB_Lehr_Speed_HMI".tHMR.dMode := "FB_LehrSpeed_IDB".tHMR.dMode;
       "DB_Lehr_Speed_HMI".tHMR.dRequestSpeedSource := "FB_LehrSpeed_IDB".tHMR.dRequestSpeedSource;

       //Move LEHR SPEED HMW
       "FB_LehrSpeed_IDB".tHMW.xAutoModeReq :=  "DB_Lehr_Speed_HMI".tHMW.xAutoModeReq;
       "FB_LehrSpeed_IDB".tHMW.xManModeReq := "DB_Lehr_Speed_HMI".tHMW.xManModeReq;
       "FB_LehrSpeed_IDB".tHMW.dManualSpeedValue_mm_min := "DB_Lehr_Speed_HMI".tHMW.dManualSpeedValue_mm_min;
       "FB_LehrSpeed_IDB".tHMW.dSpeedOverride_permil := "DB_Lehr_Speed_HMI".tHMW.dSpeedOverride_permil;
       "FB_LehrSpeed_IDB".tHMW.dSpeedSelection := "DB_Lehr_Speed_HMI".tHMW.dSpeedSelection;

      //Move LEHR SPEED ALM
       "DB_Lehr_Speed_HMI".tALM.tF := "FB_LehrSpeed_IDB".tALM.tF;
       "DB_Lehr_Speed_HMI".tALM.tS := "FB_LehrSpeed_IDB".tALM.tS;
       "DB_Lehr_Speed_HMI".tALM.tW := "FB_LehrSpeed_IDB".tALM.tW;

       //Move M203 HMR
       "DB_EmXcut_M203_SnapM201_HMI".tHMR.dDistanceSnaproll_cmm := "FB_IO_EmergencyCuttingBridge_DB".tHMR.dDistanceFromSnaproll_cmm;
       "DB_EmXcut_M203_SnapM201_HMI".tHMR.dState := "FB_IO_EmergencyCuttingBridge_DB".tHMR.dState;

       //Move M203 HMW
       "FB_IO_EmergencyCuttingBridge_DB".tHMW.xUpdateDistSnap := "DB_EmXcut_M203_SnapM201_HMI".tHMW.xUpdateDistanceSnaproll;

       "FB_IO_EmergencyCuttingBridge_DB".tHMW.dDistanceFromSnaproll_cmm := "DB_EmXcut_M203_SnapM201_HMI".tHMW.dDistanceSnaproll_cmm;
       "FB_IO_EmergencyCuttingBridge_DB".tHMW.dSnapDuration_ms := "DB_EmXcut_M203_SnapM201_HMI".tHMW.dSnapDuration_ms;
       "FB_IO_EmergencyCuttingBridge_DB".tHMW.dAccelerationDelay_ms := "DB_EmXcut_M203_SnapM201_HMI".tHMW.AccelerationDelay_ms  ;
       "FB_IO_EmergencyCuttingBridge_DB".tHMW.rBreakPosOffset_mm := "DB_EmXcut_M203_SnapM201_HMI".tHMW.rBreakPosOffset_mm;
       "FB_IO_EmergencyCuttingBridge_DB".tHMW.rPlateLenght_mm := "DB_EmXcut_M203_SnapM201_HMI".tHMW.rPlateLenght_mm;

       //Move M203 ALM 
       "DB_EmXcut_M203_SnapM201_HMI".tALM.tF :="FB_IO_EmergencyCuttingBridge_DB".tALM.tF;


       //Move OPT Manager HMR
       "DB_OPT_Manager_HMI".tHMR.dDecisionLinePosition_cmm :="FB_OptManager_V1_00_IDB".tHMR.dDecisionLinePosition_cmm;
       "DB_OPT_Manager_HMI".tHMR.dLastOptLinePosition_cmm := "FB_OptManager_V1_00_IDB".tHMR.dLastOptLinePosition_cmm;
       "DB_OPT_Manager_HMI".tHMR.dSelOptimizer := "FB_OptManager_V1_00_IDB".tHMR.dSelOptimizer;

       "DB_OPT_Manager_HMI".tHMR.dCameraGrossWander_cmm := "FB_OptManager_V1_00_IDB".tHMR.rgtRibbonData[0].dGrossWander_cmm;
       "DB_OPT_Manager_HMI".tHMR.dCameraNetWander_cmm := "FB_OptManager_V1_00_IDB".tHMR.rgtRibbonData[0].dNetWander_cmm;
       "DB_OPT_Manager_HMI".tHMR.dCameraGrossWidth_cmm:= "FB_OptManager_V1_00_IDB".tHMR.rgtRibbonData[0].dGrossWidth_cmm;
       "DB_OPT_Manager_HMI".tHMR.dCameraNetWidth_cmm := "FB_OptManager_V1_00_IDB".tHMR.rgtRibbonData[0].dNetWidth_cmm;

       "DB_OPT_Manager_HMI".tHMR.dScannerGrossWander_cmm := "FB_OptManager_V1_00_IDB".tHMR.rgtRibbonData[1].dGrossWander_cmm;
       "DB_OPT_Manager_HMI".tHMR.dScannerNetWander_cmm := "FB_OptManager_V1_00_IDB".tHMR.rgtRibbonData[1].dNetWander_cmm;
       "DB_OPT_Manager_HMI".tHMR.dScannerGrossWidth_cmm := "FB_OptManager_V1_00_IDB".tHMR.rgtRibbonData[1].dGrossWidth_cmm;
       "DB_OPT_Manager_HMI".tHMR.dScannerNetWidth_cmm := "FB_OptManager_V1_00_IDB".tHMR.rgtRibbonData[1].dNetWidth_cmm;

       //Move OPT Manager HMW
       //
       "FB_OptManager_V1_00_IDB".tHMW.xSelectOptimizerA := "DB_OPT_Manager_HMI".tHMW.xSelectOptimizerA;
       "FB_OptManager_V1_00_IDB".tHMW.xSelectOptimizerB := "DB_OPT_Manager_HMI".tHMW.xSelectOptimizerB;
       "FB_OptManager_V1_00_IDB".tHMW.xUpdateDecisionLine := "DB_OPT_Manager_HMI".tHMW.xUpdateDecisionLine;
       "FB_OptManager_V1_00_IDB".tHMW.xUpdateLastOptimizerLine := "DB_OPT_Manager_HMI".tHMW.xUpdateLastOptimizerLine;

       "FB_OptManager_V1_00_IDB".tHMW.dDecisionLinePosition_cmm := "DB_OPT_Manager_HMI".tHMW.dDecisionLinePosition_cmm;
       "FB_OptManager_V1_00_IDB".tHMW.dLastOptLinePosition_cmm := "DB_OPT_Manager_HMI".tHMW.dLastOptLinePosition_cmm;
       "FB_OptManager_V1_00_IDB".tHMW.dManualGrossWidth_cmm := "DB_OPT_Manager_HMI".tHMW.dManualGrossWidth_cmm;
       "FB_OptManager_V1_00_IDB".tHMW.dManualNetWidth_cmm := "DB_OPT_Manager_HMI".tHMW.dManualNetWidth_cmm;
       "FB_OptManager_V1_00_IDB".tHMW.dManualWander_cmm := "DB_OPT_Manager_HMI".tHMW.dManualWander_cmm;
       "FB_OptManager_V1_00_IDB".tHMW.dSelectRibbonDataSource := "DB_OPT_Manager_HMI".tHMW.dSelectRibbonDataSource;
       "FB_OptManager_V1_00_IDB".tHMW.dSelectWanderDataSource := "DB_OPT_Manager_HMI".tHMW.dSelectWanderDataSource;
       "FB_OptManager_V1_00_IDB".tHMW.dSelectWanderMode := "DB_OPT_Manager_HMI".tHMW.dSelectWanderMode;
       "FB_OptManager_V1_00_IDB".tHMW.dWanderOffset_cmm := "DB_OPT_Manager_HMI".tHMW.dWanderOffset_cmm;
       "FB_OptManager_V1_00_IDB".tHMW.dWanderRecThr_cmm := "DB_OPT_Manager_HMI".tHMW.dWanderRecThr_cmm;




       //Move SnapRoll M221 HMR
       "DB_SnapRoll_221_HMI".tHMR.xManualCommandEnabled := "FB_Snaproll_V1_00_IDB".tHMR.xManComEnSnap;

       "DB_SnapRoll_221_HMI".tHMR.tManCmd.xContrastActivation := "FB_Snaproll_V1_00_IDB".tHMR.tManCmd.xContrastActivation;
       "DB_SnapRoll_221_HMI".tHMR.tManCmd.xUp := "FB_Snaproll_V1_00_IDB".tHMR.tManCmd.xUp;

       "DB_SnapRoll_221_HMI".tHMR.dStatus := "FB_Snaproll_V1_00_IDB".tHMR.dStatus;


       //Move SnapRoll M221  HMW
       "FB_Snaproll_V1_00_IDB".tHMW.xEnDisManComSnap :="DB_SnapRoll_221_HMI".tHMW.xEnableManualCommand ;
       "FB_Snaproll_V1_00_IDB".tHMW.tMan.xContrastActivation :="DB_SnapRoll_221_HMI".tHMW.tManCmd.xContrastActivation ;
       "FB_Snaproll_V1_00_IDB".tHMW.tMan.xUp :="DB_SnapRoll_221_HMI".tHMW.tManCmd.xUp ;
       "FB_Snaproll_V1_00_IDB".tHMW.dMaxPlateLenghtEnableContrast_cmm :="DB_SnapRoll_221_HMI".tHMW.dMaxPlateLenghtEnableContrast_cmm;
       "FB_Snaproll_V1_00_IDB".tHMW.dOffsetSnap_cmm :="DB_SnapRoll_221_HMI".tHMW.dOffsetSnap_cmm ;
       "FB_Snaproll_V1_00_IDB".tHMW.dReactTime_ms :="DB_SnapRoll_221_HMI".tHMW.dReactTime_ms ;
       "FB_Snaproll_V1_00_IDB".tHMW.dTimeUp_ms :="DB_SnapRoll_221_HMI".tHMW.dTimeUp_ms ;


       //Move SnapRoll M221 ALM  
       "DB_SnapRoll_221_HMI".tALM.tF :="FB_Snaproll_V1_00_IDB".tALM.tF ;
       "DB_SnapRoll_221_HMI".tALM.tS :="FB_Snaproll_V1_00_IDB".tALM.tS ;
       "DB_SnapRoll_221_HMI".tALM.tW :="FB_Snaproll_V1_00_IDB".tALM.tW ;

       //Move DIGITIZER PH   HMR 
       "DB_Digitizer_Break_detector_HMI".tHMR."xPhotoStatus[0]"  :="FB_BD_DigitizerPH_V1_00_IDB".tHMR.rgxPhotoStatus[0];
       "DB_Digitizer_Break_detector_HMI".tHMR."xPhotoStatus[1]" := "FB_BD_DigitizerPH_V1_00_IDB".tHMR.rgxPhotoStatus[1];

       "DB_Digitizer_Break_detector_HMI".tHMR.dDistanceSnaproll_cmm := "FB_BD_DigitizerPH_V1_00_IDB".tHMR.dDistanceSnaproll_cmm;
       "DB_Digitizer_Break_detector_HMI".tHMR.dStatus := "FB_BD_DigitizerPH_V1_00_IDB".tHMR.dStatus;
       "DB_Digitizer_Break_detector_HMI".tHMR."dPhotoAbilitation[0]" := "FB_BD_DigitizerPH_V1_00_IDB".tHMR.rgdPhotoAbilitation[0];
       "DB_Digitizer_Break_detector_HMI".tHMR."dPhotoAbilitation[1]" := "FB_BD_DigitizerPH_V1_00_IDB".tHMR.rgdPhotoAbilitation[1];

       //Move DIGITIZER PH   HMW
       "FB_BD_DigitizerPH_V1_00_IDB".tHMW.xUpdateDistanceSnap := "DB_Digitizer_Break_detector_HMI".tHMW.xUpdateDistanceSnaproll;
       "FB_BD_DigitizerPH_V1_00_IDB".tHMW.rgxEnabledPhotocell[0] :="DB_Digitizer_Break_detector_HMI".tHMW."xPhotoEnabled[0]";
       "FB_BD_DigitizerPH_V1_00_IDB".tHMW.rgxEnabledPhotocell[1] :="DB_Digitizer_Break_detector_HMI".tHMW."xPhotoEnabled[0]";
       "FB_BD_DigitizerPH_V1_00_IDB".tHMW.dDistanceSnaproll_cmm := "DB_Digitizer_Break_detector_HMI".tHMW.dDistanceSnaproll_cmm;
       "FB_BD_DigitizerPH_V1_00_IDB".tHMW.dMinBreakSize_cmm := "DB_Digitizer_Break_detector_HMI".tHMW.dMinBreakSize_cmm;

       //Move DIGITIZER PH   ALM
       "DB_Digitizer_Break_detector_HMI".tALM.tF := "FB_BD_DigitizerPH_V1_00_IDB".tALM.tF;
       "DB_Digitizer_Break_detector_HMI".tALM.tS := "FB_BD_DigitizerPH_V1_00_IDB".tALM.tS;
       "DB_Digitizer_Break_detector_HMI".tALM.tW := "FB_BD_DigitizerPH_V1_00_IDB".tALM.tW;


       //Move CROSS CUT OPT HMR  
       "DB_CrossCut_Opt_HMI".tHMR.xEnabledPriority := "FB_CrossCut_Opt_V1_00_IDB".tHMR.xEnabledPriority;

       //Move CROSS CUT OPT HMW 
       "FB_CrossCut_Opt_V1_00_IDB".tHMW.xEnDisPriority:= "DB_CrossCut_Opt_HMI".tHMW.xEnDisPriority;

       //Move CROSS CUT #1 HMR 

